               REGION "BUTTON 3"
                   #btnActivateInt[3] := #btn3Activate;
                   #btnModeInt[3] := #btn3Mode;
                   #btnGroup[3] := #btn3Group;
                   #btnClrOn1Int[3] := #btn3ColorOn1;
                   #btnClrOn2Int[3] := #btn3ColorOn2;
                   #btnClrOffInt[3] := #btn3ColorOff;
               END_REGION

               REGION "BUTTON 4"
                   #btnActivateInt[4] := #btn4Activate;
                   #btnModeInt[4] := #btn4Mode;
                   #btnGroup[4] := #btn4Group;
                   #btnClrOn1Int[4] := #btn4ColorOn1;
                   #btnClrOn2Int[4] := #btn4ColorOn2;
                   #btnClrOffInt[4] := #btn4ColorOff;
               END_REGION

               REGION "BUTTON 5"
                   #btnActivateInt[5] := #btn5Activate;
                   #btnModeInt[5] := #btn5Mode;
                   #btnGroup[5] := #btn5Group;
                   #btnClrOn1Int[5] := #btn5ColorOn1;
                   #btnClrOn2Int[5] := #btn5ColorOn2;
                   #btnClrOffInt[5] := #btn5ColorOff;
               END_REGION

               REGION "BUTTON 6"
                   #btnActivateInt[6] := #btn6Activate;
                   #btnModeInt[6] := #btn6Mode;
                   #btnGroup[6] := #btn6Group;
                   #btnClrOn1Int[6] := #btn6ColorOn1;
                   #btnClrOn2Int[6] := #btn6ColorOn2;
                   #btnClrOffInt[6] := #btn6ColorOff;
               END_REGION

               REGION "BUTTON 7"
                   #btnActivateInt[7] := #btn7Activate;
                   #btnModeInt[7] := #btn7Mode;
                   #btnGroup[7] := #btn7Group;
                   #btnClrOn1Int[7] := #btn7ColorOn1;
                   #btnClrOn2Int[7] := #btn7ColorOn2;
                   #btnClrOffInt[7] := #btn7ColorOff;
               END_REGION

           END_REGION

           REGION "RECOLOR BUTTON MASKS"
               FOR #i1 := 0 TO 7 DO

                   REGION "ON COLOR 1"
                       IF (#btnClrOn1Int[#i1] = 'red') THEN
                           #btnClrMskOn1Int[#i1] := SHL(IN := #btnMskRed, N := INT_TO_ULINT(#i1));
                       ELSIF (#btnClrOn1Int[#i1] = 'green') THEN
                           #btnClrMskOn1Int[#i1] := SHL(IN := #btnMskGreen, N := INT_TO_ULINT(#i1));
                       ELSIF (#btnClrOn1Int[#i1] = 'blue') THEN
                           #btnClrMskOn1Int[#i1] := SHL(IN := #btnMskBlue, N := INT_TO_ULINT(#i1));
                       ELSIF (#btnClrOn1Int[#i1] = 'yellow') THEN
                           #btnClrMskOn1Int[#i1] := SHL(IN := #btnMskYellow, N := INT_TO_ULINT(#i1));
                       ELSIF (#btnClrOn1Int[#i1] = 'white') THEN
                           #btnClrMskOn1Int[#i1] := SHL(IN := #btnMskWhite, N := INT_TO_ULINT(#i1));
                       ELSIF (#btnClrOn1Int[#i1] = 'off') THEN
                           #btnClrMskOn1Int[#i1] := 0;
                       END_IF;
                   END_REGION

                   REGION "ON COLOR 2"
                       IF (#btnClrOn2Int[#i1] = 'red') THEN
                           #btnClrMskOn2Int[#i1] := SHL(IN := #btnMskRed, N := INT_TO_ULINT(#i1));
                       ELSIF (#btnClrOn2Int[#i1] = 'green') THEN
                           #btnClrMskOn2Int[#i1] := SHL(IN := #btnMskGreen, N := INT_TO_ULINT(#i1));
                       ELSIF (#btnClrOn2Int[#i1] = 'blue') THEN
                           #btnClrMskOn2Int[#i1] := SHL(IN := #btnMskBlue, N := INT_TO_ULINT(#i1));
                       ELSIF (#btnClrOn2Int[#i1] = 'yellow') THEN
                           #btnClrMskOn2Int[#i1] := SHL(IN := #btnMskYellow, N := INT_TO_ULINT(#i1));
                       ELSIF (#btnClrOn2Int[#i1] = 'white') THEN
                           #btnClrMskOn2Int[#i1] := SHL(IN := #btnMskWhite, N := INT_TO_ULINT(#i1));
                       ELSIF (#btnClrOn2Int[#i1] = 'off') THEN
                           #btnClrMskOn2Int[#i1] := 0;
                       END_IF;
                   END_REGION

                   REGION "OFF COLOR"
                       IF (#btnClrOffInt[#i1] = 'red') THEN
                           #btnClrMskOffInt[#i1] := SHL(IN := #btnMskRed, N := INT_TO_ULINT(#i1));
                       ELSIF (#btnClrOffInt[#i1] = 'green') THEN
                           #btnClrMskOffInt[#i1] := SHL(IN := #btnMskGreen, N := INT_TO_ULINT(#i1));
                       ELSIF (#btnClrOffInt[#i1] = 'blue') THEN
                           #btnClrMskOffInt[#i1] := SHL(IN := #btnMskBlue, N := INT_TO_ULINT(#i1));
                       ELSIF (#btnClrOffInt[#i1] = 'yellow') THEN
                           #btnClrMskOffInt[#i1] := SHL(IN := #btnMskYellow, N := INT_TO_ULINT(#i1));
                       ELSIF (#btnClrOffInt[#i1] = 'white') THEN
                           #btnClrMskOffInt[#i1] := SHL(IN := #btnMskWhite, N := INT_TO_ULINT(#i1));
                       ELSIF (#btnClrOffInt[#i1] = 'off') THEN
                           #btnClrMskOffInt[#i1] := 0;
                       END_IF;
                   END_REGION

               END_FOR;
           END_REGION

       END_IF;
   END_REGION

   REGION "HART INIT"
       IF #hardInit THEN
           FOR #i1 := 0 TO 7 DO
               #btnStateArrayInt[#i1] := FALSE;
           END_FOR;
       END_IF;
   END_REGION


   REGION "TRANFER PARAMETERS TO ARRAYS"
       // raw pb data
       #btnInInt := #btnIn;
       // flashing modes
       #btnFlashInt[0] := #btn0Flash;
       #btnFlashInt[1] := #btn1Flash;
       #btnFlashInt[2] := #btn2Flash;
       #btnFlashInt[3] := #btn3Flash;
       #btnFlashInt[4] := #btn4Flash;
       #btnFlashInt[5] := #btn5Flash;
       #btnFlashInt[6] := #btn6Flash;
       #btnFlashInt[7] := #btn7Flash;
   END_REGION

   REGION "EVALUATE BUTTONS"
       FOR #i1 := 0 TO 7 DO

           REGION "TRANSFER BUTTON PRESSES TO ARRAY"
               #btnEval := SHR(IN := #btnInInt, N := INT_TO_ULINT(#i1));
               #btnInArrayNew[#i1] := #btnEval.%X0;
               #btnEval := b#16#0;
           END_REGION

           REGION "SET BUTTON STATE"

               REGION "BUTTON ACTIVE"
                   IF #btnActivateInt[#i1] THEN

                       REGION "MAINTAINED"
                           IF #btnModeInt[#i1] THEN

                               REGION "RISING EDGE OF PRESS"
                                   IF #btnInArrayNew[#i1] AND NOT #btnInArrayOld[#i1] THEN

                                       REGION "CHECK FOR GROUP MEMBERSHIP"
                                           FOR #i2 := 0 TO 7 DO

                                               REGION "NOT IN NULL GROUP"
                                                   IF (#btnGroup[#i2] <> 0) THEN

                                                       REGION "SKIP SELF"
                                                           IF (#i2 <> #i1) THEN

                                                               REGION "GROUPS MATCH"
                                                                   IF #btnGroup[#i1] = #btnGroup[#i2] THEN
                                                                       REGION "DEACTIVATE OTHER GROUP MEMBERS"
                                                                           #btnStateArrayInt[#i2] := FALSE;
                                                                       END_REGION

                                                                   END_IF;
                                                               END_REGION

                                                           END_IF;
                                                       END_REGION

                                                   END_IF;
                                               END_REGION

                                           END_FOR;
                                       END_REGION

                                       REGION "TOGGLE STATE"
                                           #btnStateArrayInt[#i1] := NOT #btnStateArrayInt[#i1];
                                       END_REGION

                                   END_IF;
                               END_REGION

                           END_IF;
                       END_REGION

                       REGION "MOMENTARY"
                           IF NOT #btnModeInt[#i1] THEN
                               #btnStateArrayInt[#i1] := #btnInArrayNew[#i1];
                           END_IF;
                       END_REGION

                   END_IF;
               END_REGION

               REGION "BUTTON INACTIVE"
                   IF NOT #btnActivateInt[#i1] THEN
                       #btnStateArrayInt[#i1] := FALSE;
                   END_IF;
               END_REGION

           END_REGION

           REGION "ANIMATE BUTTONS"

               REGION "BUTTON ON FLASH BIT OFF"
                   IF #btnStateArrayInt[#i1] AND NOT #btnFlashInt[#i1] THEN
                       #btnColors := #btnColors AND ROL(IN := #btnMskBlack, N := INT_TO_ULINT(#i1));
                       #btnColors := #btnColors OR #btnClrMskOn1Int[#i1];
                   END_IF;
               END_REGION

               REGION "BUTTON ON FLASH BIT ON"
                   IF #btnStateArrayInt[#i1] AND #btnFlashInt[#i1] THEN
                       #btnColors := #btnColors AND ROL(IN := #btnMskBlack, N := INT_TO_ULINT(#i1));
                       #btnColors := #btnColors OR #btnClrMskOn2Int[#i1];
                   END_IF;
               END_REGION

               REGION "BUTTON OFF"
                   IF NOT #btnStateArrayInt[#i1] THEN
                       #btnColors := #btnColors AND ROL(IN := #btnMskBlack, N := INT_TO_ULINT(#i1));
                       #btnColors := #btnColors OR #btnClrMskOffInt[#i1];
                   END_IF;
               END_REGION

           END_REGION

       END_FOR;
   END_REGION

   REGION "CHANGE DETECTION"
       #btnInArrayOld := #btnInArrayNew;
   END_REGION

   REGION "OUTPUT"
       #btnColorsOut := #btnColors;
       #btnStatesOut := #btnStateArrayInt;
   END_REGION
END_FUNCTION_BLOCK

FUNCTION "Physical to Global" : Void   // FC1, LAD
{ S7_Optimized_Access := 'TRUE' }
VERSION : 0.1
   VAR_IN_OUT
      stations : "Stations";
   END_VAR
   VAR_TEMP
      i : Int;
      kp8In : DWord;
   END_VAR
BEGIN

REGION Network 1 (SCL): MAIN LOOP
   FOR #i := 0 TO "stnCount" DO

       CASE #i OF
           "VOLVO 16 01":
               #kp8In := "VOLVO 16 01 KP8 In";
           "VOLVO 16 02":
               #kp8In := "VOLVO 16 02 KP8 In";
           "VOLVO 16 03":
               #kp8In := "VOLVO 16 03 KP8 In";
           "VOLVO 16 04":
               #kp8In := "VOLVO 16 04 KP8 In";
           "VOLVO 16 05":
               #kp8In := "VOLVO 16 05 KP8 In";
           "VOLVO 16 06":
               #kp8In := "VOLVO 16 06 KP8 In";
           "VOLVO 16 07":
               #kp8In := "VOLVO 16 07 KP8 In";
           "VOLVO 16 08":
               #kp8In := "VOLVO 16 08 KP8 In";
           "VOLVO 16 09":
               #kp8In := "VOLVO 16 09 KP8 In";
           "VOLVO 16 10":
               #kp8In := "VOLVO 16 10 KP8 In";
           "VOLVO 16 11":
               #kp8In := "VOLVO 16 11 KP8 In";
           "CHM 01":
               #kp8In := "CHM 01 KP8 In";
           "CHM 02":
               #kp8In := "CHM 02 KP8 In";
           "CHM 03":
               #kp8In := "CHM 03 KP8 In";
           "CHM 04":
               #kp8In := "CHM 04 KP8 In";
           "CHM 05":
               #kp8In := "CHM 05 KP8 In";
           "CDO 01":
               #kp8In := "CDO 01 KP8 In";
           "CDO 02":
               #kp8In := "CDO 02 KP8 In";
           "CDO 03":
               #kp8In := "CDO 03 KP8 In";
           "BFL 01":
               #kp8In := "BFL 01 KP8 In";
           "BFL 02":
               #kp8In := "BFL 02 KP8 In";
           "BFL 03":
               #kp8In := "BFL 03 KP8 In";
           "LGS 01":
               #kp8In := "LGS 01 KP8 In";
           "LGS 02":
               #kp8In := "LGS 02 KP8 In";

       END_CASE;

       #stations.me[#i].kp8In := #kp8In.%B3;

   END_FOR;
END_REGION
END_FUNCTION

FUNCTION "Time to WString" : WString   // FC2, SCL
{ S7_Optimized_Access := 'TRUE' }
VERSION : 0.1
   VAR_INPUT
      "Time" : Time;
   END_VAR
   VAR_TEMP
      "Time as DInt" : DInt;
      "Hours 10s Place" : DInt;
      "Hours 1s Place" : DInt;
      "Minutes 10s Place" : DInt;
      "Minutes 1s Place" : DInt;
      "Seconds 10s Place" : DInt;
      "Seconds 1s Place" : DInt;
      "Time Elements" : Array[0..4] of WString;
      Length : Int;
      "String Box" : WString;
      "DInt Box" : DInt;
   END_VAR
   VAR CONSTANT
      "Milliseconds per 10 Hours" : DInt := 36000000;
      "Milliseconds per Hour" : DInt := 3600000;
      "Milliseconds per 10 Minutes" : DInt := 600000;
      "Milliseconds per Minute" : DInt := 60000;
      "Milliseconds per 10 Seconds" : DInt := 10000;
      "Milliseconds per Second" : DInt := 1000;
   END_VAR
BEGIN
   REGION GET INPUT
       #"Time as DInt" := #Time;
   END_REGION

   REGION CONVERT TIME INTO INDIVIDUAL PLACE VALUES
       #"Minutes 10s Place" := #"Time as DInt" / #"Milliseconds per 10 Minutes";
       #"Minutes 1s Place" := (#"Time as DInt" / #"Milliseconds per Minute") MOD 10;
       #"Seconds 10s Place" := (#"Time as DInt" MOD #"Milliseconds per Minute") / #"Milliseconds per 10 Seconds";
       #"Seconds 1s Place" := (#"Time as DInt" / #"Milliseconds per Second") MOD 10;
   END_REGION

   REGION "ADD SIGN"
       #"Time Elements"[0] := wstring#'';
       IF #"Minutes 10s Place" < 0 OR
           #"Minutes 1s Place" < 0 OR
           #"Seconds 10s Place" < 0 OR
           #"Seconds 1s Place" < 0 THEN
            #"Time Elements"[0] := wstring#'-';
       END_IF;
   END_REGION

   REGION CONVERT PLACE VALUES INTO COMPONENT STRINGS
       // MINUTES
       #"DInt Box" := #"Minutes 10s Place" * 10 + #"Minutes 1s Place";
       #"String Box" := DINT_TO_WSTRING(IN := #"DInt Box");
       #"String Box" := "Strip Sign"("WString":=#"String Box");
       #"String Box" := "Add Leading"("Leading Character" := WCHAR#'0',
                                      "Desired Length" := 2,
                                      "String" := #"String Box");
       #"Time Elements"[1] := #"String Box";
       // COLON
       #"Time Elements"[2] := WSTRING#':';
       // SECONDS
       #"DInt Box" := #"Seconds 10s Place" * 10 + #"Seconds 1s Place";
       #"String Box" := DINT_TO_WSTRING(IN := #"DInt Box");
       #"String Box" := "Strip Sign"("WString":=#"String Box");
       #"String Box" := "Add Leading"("Leading Character" := WCHAR#'0',
                                      "Desired Length" := 2,
                                      "String" := #"String Box");
       #"Time Elements"[3] := #"String Box";
   END_REGION


   REGION RETURN VALUE
       #"Time to WString" := CONCAT_WSTRING(IN1 := #"Time Elements"[0],
                                            IN2 := #"Time Elements"[1],
                                            IN3 := #"Time Elements"[2],
                                            IN4 := #"Time Elements"[3]);
   END_REGION
END_FUNCTION

FUNCTION "Strip Sign" : WString   // FC3, SCL
{ S7_Optimized_Access := 'TRUE' }
VERSION : 0.1
   VAR_INPUT
      WString : WString;
   END_VAR
   VAR_TEMP
      Length : Int;
      "String Box" : WString;
      "Test Character" : WString;
   END_VAR
   VAR CONSTANT
      "+" : WChar := WCHAR#'+';
      "-" : WChar := WCHAR#'-';
   END_VAR
BEGIN
   #"String Box" := #WString;
   #"Test Character" := LEFT_WSTRING(IN := #"String Box",
                                     L := 1);
   IF #"Test Character" = #"+" OR #"Test Character" = #"-" THEN
       #Length := LEN(#"String Box");
       #"String Box" := RIGHT_WSTRING(IN := #"String Box", L := #Length - 1);

   END_IF;
   #"Strip Sign" := #"String Box";
END_FUNCTION

FUNCTION "Add Leading" : WString   // FC4, SCL
{ S7_Optimized_Access := 'TRUE' }
VERSION : 0.1
   VAR_INPUT
      "Leading Character" : WChar;
      "Desired Length" : USInt;
      "String" : WString;
   END_VAR
   VAR_TEMP
      Length : Int;
      "String Box" : WString;
      Constant : WString;
   END_VAR
BEGIN
   #"String Box" := #String;
   #Length := LEN(#"String Box");

   WHILE #Length < #"Desired Length" DO
       #"String Box" := CONCAT_WSTRING(IN1 := #"Leading Character",
                                       IN2 := #"String Box");
       #Length := LEN(#"String Box");
   END_WHILE;

   #"Add Leading" := #"String Box";
END_FUNCTION

FUNCTION "Global to Physical" : Void   // FC5, LAD
{ S7_Optimized_Access := 'TRUE' }
VERSION : 0.1
   VAR_IN_OUT
      stations : "Stations";
   END_VAR
   VAR_TEMP
      i : Int;
      j : Int;
      IO : DWord;
      "KP8 In" : DWord;
      "KP8 Out" : DWord;
      Card : Int;
      stnCount : Int;
   END_VAR
   VAR CONSTANT
      "VOLVO 16 01" : Int := 0;
      "VOLVO 16 02" : Int := 1;
      "VOLVO 16 03" : Int := 2;
      "VOLVO 16 04" : Int := 3;
      "VOLVO 16 05" : Int := 4;
      "VOLVO 16 06" : Int := 5;
      "VOLVO 16 07" : Int := 6;
      "VOLVO 16 08" : Int := 7;
      "VOLVO 16 09" : Int := 8;
      "VOLVO 16 10" : Int := 9;
      "VOLVO 16 11" : Int := 10;
      "CHM 01" : Int := 11;
      "CHM 02" : Int := 12;
      "CHM 03" : Int := 13;
      "CHM 04" : Int := 14;
      "CHM 05" : Int := 15;
      "CDO 01" : Int := 16;
      "CDO 02" : Int := 17;
      "CDO 03" : Int := 18;
      "BFL 01" : Int := 19;
      "BFL 02" : Int := 20;
      "BFL 03" : Int := 21;
      "LGS 01" : Int := 22;
      "LGS 02" : Int := 23;
   END_VAR
BEGIN

REGION Network 1: ARRAY LIMIT FOR STATION COUNT
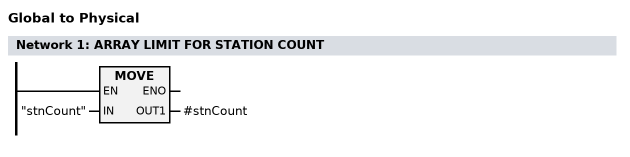
   RUNG wire#powerrail
      Move(in := "stnCount", out1 => #stnCount)
   END_RUNG
   // the same network as SCL:
   #stnCount := "stnCount";
END_REGION

REGION Network 2 (SCL): MAIN LOOP
   FOR #i := 0 TO #stnCount DO

       #IO := #stations.me[#i].stackLightOut;
       #"KP8 Out" := #stations.me[#i].kp8Out;

       CASE #i OF
           #"VOLVO 16 01":
               "VOLVO 16 01 IO" := #IO;
               "VOLVO 16 01 KP8 Out" := #"KP8 Out";
           #"VOLVO 16 02":
               "VOLVO 16 02 IO" := #IO;
               "VOLVO 16 02 KP8 Out" := #"KP8 Out";
           #"VOLVO 16 03":
               "VOLVO 16 03 IO" := #IO;
               "VOLVO 16 03 KP8 Out" := #"KP8 Out";
           #"VOLVO 16 04":
               "VOLVO 16 04 IO" := #IO;
               "VOLVO 16 04 KP8 Out" := #"KP8 Out";
           #"VOLVO 16 05":
               "VOLVO 16 05 IO" := #IO;
               "VOLVO 16 05 KP8 Out" := #"KP8 Out";
           #"VOLVO 16 06":
               "VOLVO 16 06 IO" := #IO;
               "VOLVO 16 06 KP8 Out" := #"KP8 Out";
           #"VOLVO 16 07":
               "VOLVO 16 07 IO" := #IO;
               "VOLVO 16 07 KP8 Out" := #"KP8 Out";
           #"VOLVO 16 08":
               "VOLVO 16 08 IO" := #IO;
               "VOLVO 16 08 KP8 Out" := #"KP8 Out";
           #"VOLVO 16 09":
               "VOLVO 16 09 IO" := #IO;
               "VOLVO 16 09 KP8 Out" := #"KP8 Out";
           #"VOLVO 16 10":
               "VOLVO 16 10 IO" := #IO;
               "VOLVO 16 10 KP8 Out" := #"KP8 Out";
           #"VOLVO 16 11":
               "VOLVO 16 11 IO" := #IO;
               "VOLVO 16 11 KP8 Out" := #"KP8 Out";
           #"CHM 01":
               "CHM 01 IO" := #IO;
               "CHM 01 KP8 Out" := #"KP8 Out";
           #"CHM 02":
               "CHM 02 IO" := #IO;
               "CHM 02 KP8 Out" := #"KP8 Out";
           #"CHM 03":
               "CHM 03 IO" := #IO;
               "CHM 03 KP8 Out" := #"KP8 Out";
           #"CHM 04":
               "CHM 04 IO" := #IO;
               "CHM 04 KP8 Out" := #"KP8 Out";
           #"CHM 05":
               "CHM 05 IO" := #IO;
               "CHM 05 KP8 Out" := #"KP8 Out";
           #"CDO 01":
               "CDO 01 IO" := #IO;
               "CDO 01 KP8 Out" := #"KP8 Out";
           #"CDO 02":
               "CDO 02 IO" := #IO;
               "CDO 02 KP8 Out" := #"KP8 Out";
           #"CDO 03":
               "CDO 03 IO" := #IO;
               "CDO 03 KP8 Out" := #"KP8 Out";
           #"BFL 01":
               "BFL 01 IO" := #IO;
               "BFL 01 KP8 Out" := #"KP8 Out";
           #"BFL 02":
               "BFL 02 IO" := #IO;
               "BFL 02 KP8 Out" := #"KP8 Out";
           #"BFL 03":
               "BFL 03 IO" := #IO;
               "BFL 03 KP8 Out" := #"KP8 Out";
           #"LGS 01":
               "LGS 01 IO" := #IO;
               "LGS 01 KP8 Out" := #"KP8 Out";
           #"LGS 02":
               "LGS 02 IO" := #IO;
               "LGS 02 KP8 Out" := #"KP8 Out";

       END_CASE;

   END_FOR;
END_REGION
END_FUNCTION

FUNCTION "Select Stations" : Void   // FC6, SCL
{ S7_Optimized_Access := 'TRUE' }
VERSION : 0.1
   VAR_INPUT
      mode : Bool;   // TRUE = select; FALSE = deselect
   END_VAR
   VAR_IN_OUT
      stations : "Stations";
   END_VAR
   VAR_TEMP
      i : Int;
      stnCount : Int;
   END_VAR
   VAR CONSTANT
      stationCount : Int := 22;
   END_VAR
BEGIN
   REGION "GET STATION COUNT"
       #stnCount := "stnCount";
   END_REGION

   REGION "SELECT STATIONS"
       FOR #i := 0 TO #stnCount DO
           #stations.me[#i].settings.selected := #mode;
       END_FOR;
   END_REGION
END_FUNCTION

FUNCTION "Dark Mode" : Void   // FC7, SCL
{ S7_Optimized_Access := 'TRUE' }
VERSION : 0.1
   VAR_IN_OUT
      animate : USInt;
   END_VAR
   VAR_TEMP
      ani : USInt;
   END_VAR
   VAR CONSTANT
      redFlashing : USInt := 12;
      invisible : USInt := 255;
      darkMode : USInt := 1;
      disabled : USInt := 254;
   END_VAR
BEGIN
   REGION "COPY TO LOCAL"
       #ani := #animate;
   END_REGION


   REGION "APPLY DARK MODE"
       CASE #ani OF
           #redFlashing, #invisible, 0, #disabled:
               #ani := #ani;
           ELSE
               #ani += #darkMode;
       END_CASE;
   END_REGION


   REGION "OUTPUT"
       #animate := #ani;
   END_REGION
END_FUNCTION

FUNCTION "Select Buttons" : Void   // FC8, SCL
{ S7_Optimized_Access := 'TRUE' }
VERSION : 0.1
   VAR_INPUT
      mode : Bool;   // TRUE = select; FALSE = deselect
   END_VAR
   VAR_IN_OUT
      stations : "Stations";
   END_VAR
   VAR_TEMP
      btnCount : Int;
      i : Int;
      j : Int;
      selected : Bool;
      stnCount : Int;
   END_VAR
   VAR CONSTANT
      buttonCount : Int := 5;
   END_VAR
BEGIN
   REGION "COPY TO LOCAL"
       #btnCount := "ptsPerStn";
       #stnCount := "stnCount";
   END_REGION

   REGION "SELECT BUTTONS"
       FOR #i := 0 TO #stnCount DO

           REGION "SELCT ALL BUTTONS ON SELECTED STATION"
               #selected := #stations.me[#i].settings.selected;
               IF #selected THEN

                   REGION "LOOP THROUGH BUTTONS"
                       FOR #j := 0 TO #btnCount DO
                           #stations.me[#i].settings.btnSelection[#j] := #mode;
                       END_FOR;
                   END_REGION

               END_IF;
           END_REGION

       END_FOR;
   END_REGION
END_FUNCTION

FUNCTION "Animate Bool" : USInt   // FC9, SCL
{ S7_Optimized_Access := 'TRUE' }
VERSION : 0.1
   VAR_INPUT
      colorTrue : USInt;
      colorFalse : USInt;
      evalSignal : Bool;
   END_VAR
   VAR_TEMP
      animate : USInt;
   END_VAR
BEGIN
   REGION "FALSE COLOR"
       IF NOT #evalSignal THEN
           #animate := #colorFalse;
       END_IF;
   END_REGION

   REGION "TRUE COLOR"
       IF #evalSignal THEN
           #animate := #colorTrue;
       END_IF;
   END_REGION

   REGION "FUNCTION RETURN"
       #"Animate Bool" := #animate;
   END_REGION
END_FUNCTION

FUNCTION "WString to Time" : Time   // FC10, SCL
{ S7_Optimized_Access := 'TRUE' }
VERSION : 0.1
   VAR_INPUT
      WString : WString;
   END_VAR
   VAR_TEMP
      Count : UInt;
      "DInt Box" : DInt;
      "String Box" : WString [5];
      "Time Box" : Time;
      "WChar Array" : Array[0..4] of WChar;
   END_VAR
   VAR CONSTANT
      "ms/(10 hr)" : DInt := 36000000;
      "ms/hr" : DInt := 3600000;
      "ms/(10 min)" : DInt := 600000;
      "ms/min" : DInt := 60000;
      "ms/(10 sec)" : DInt := 10000;
      "ms/sec" : DInt := 1000;
   END_VAR
BEGIN
   REGION EXPLODE INPUT

       #"String Box" := #WString;
       IF #"String Box" = WSTRING#'' THEN
           #"String Box" := WSTRING#'00:00';
       END_IF;

       Strg_TO_Chars(Strg := #"String Box",
                     pChars := 0,
                     Cnt => #Count,
                     Chars := #"WChar Array");

   END_REGION

   REGION CONVERT ARRAY ELEMENTS TO TIME

       // 10S OF MINUTES
       #"DInt Box" := WCHAR_TO_DINT(IN := #"WChar Array"[0]) - 16#30;
       #"Time Box" := #"Time Box" + #"DInt Box" * #"ms/(10 min)";

       // MINUTES
       #"DInt Box" := WCHAR_TO_DINT(IN := #"WChar Array"[1]) - 16#30;
       #"Time Box" := #"Time Box" + #"DInt Box" * #"ms/min";

       // 10S OF SECONDS
       #"DInt Box" := WCHAR_TO_DINT(IN := #"WChar Array"[3]) - 16#30;
       #"Time Box" := #"Time Box" + #"DInt Box" * #"ms/(10 sec)";

       // SECONDS
       #"DInt Box" := WCHAR_TO_DINT(IN := #"WChar Array"[4]) - 16#30;
       #"Time Box" := #"Time Box" + #"DInt Box" * #"ms/sec";

   END_REGION


   REGION RETURN VALUE

       #"WString to Time" := #"Time Box";

   END_REGION
END_FUNCTION

FUNCTION "Get Part Call Row Number" : Int   // FC11, SCL
{ S7_Optimized_Access := 'TRUE' }
VERSION : 0.1
   VAR_IN_OUT
      partCall : "Part Call Screen";
   END_VAR
   VAR_TEMP
      hmiRows : Int;
      i : Int;
      selectedRow : Int;
   END_VAR
BEGIN
   REGION "GET NUMBER OF HMI ROWS"
       #hmiRows := "partReqHmiRowCount";
   END_REGION

   REGION "LOOP THROUGH HMI ROWS
       FOR #i := 0 TO #hmiRows DO

           REGION "FIND SELECTED ROW"
               IF #partCall.row[#i].pbSelection.actuate THEN
                   // selected row as int
                   #selectedRow := #i + 1;
                   EXIT;
               END_IF;
           END_REGION

       END_FOR;
   END_REGION

   REGION "RETURN ROW NUMBER"
       #"Get Part Call Row Number" := #selectedRow;
   END_REGION
END_FUNCTION

FUNCTION "Address to Station and Button" : Void   // FC12, SCL
{ S7_Optimized_Access := 'TRUE' }
VERSION : 0.1
   VAR_INPUT
      address : UInt;
   END_VAR
   VAR_OUTPUT
      station : UInt;
      button : UInt;
   END_VAR
BEGIN
   #station := #address / 10;
   #button := #address MOD 10;
END_FUNCTION

FUNCTION "WString Timer to Real" : Real   // FC13, SCL
{ S7_Optimized_Access := 'TRUE' }
VERSION : 0.1
   VAR_INPUT
      wstring : WString;
   END_VAR
   VAR CONSTANT
      msPerSec : Real := 1000.0;
   END_VAR
BEGIN
   #"WString Timer to Real" := DINT_TO_REAL(TIME_TO_DINT("WString to Time"(#wstring))) / #msPerSec;
END_FUNCTION

FUNCTION "Real to WString Timer" : WString   // FC14, SCL
{ S7_Optimized_Access := 'TRUE' }
VERSION : 0.1
   VAR_INPUT
      realVal : Real;
   END_VAR
   VAR CONSTANT
      msPerSec : Real := 1000.0;
   END_VAR
BEGIN
   #"Real to WString Timer" := "Time to WString"(DINT_TO_TIME(REAL_TO_DINT(#realVal * #msPerSec)));
END_FUNCTION

FUNCTION "Populate Dropzone IO Field" : WString   // FC15, SCL
{ S7_Optimized_Access := 'TRUE' }
VERSION : 0.1
   VAR_INPUT
      dzAsInt : USInt;
   END_VAR
BEGIN
   #"Populate Dropzone IO Field" := "Strip Sign"(USINT_TO_WSTRING(#dzAsInt));
END_FUNCTION

FUNCTION "Get Station Selection Number" : Void   // FC16, SCL
{ S7_Optimized_Access := 'TRUE' }
VERSION : 0.1
   VAR_INPUT
      next : Bool;   // 'next' or 'prev'
      prev : Bool;
      stations : "Stations";
   END_VAR
   VAR_IN_OUT
      selStnNumber : Int;
   END_VAR
   VAR_TEMP
      i : Int;
      stnCount : Int;
      stnSelected : Bool;
   END_VAR
BEGIN
   REGION "COPY TO LOCAL"
       #stnCount := "stnCount";
   END_REGION

   REGION "INITIALIZE INDEX"
       #i := #selStnNumber;
   END_REGION

   REGION "PREVIOUS MODE"

       REGION "DECREMENT"
           IF #prev THEN
               #i -= 1;
           END_IF;
       END_REGION

       REGION "LOW LIMIT ROLLOVER"
           IF #i < 0 THEN
               #i := #stnCount;
           END_IF;
       END_REGION

   END_REGION

   REGION "NEXT MODE"

       REGION "INCREMENT"
           IF #next THEN
               #i += 1;
           END_IF;
       END_REGION

       REGION "HIGH LIMIT ROLLOVER"
           IF #i > #stnCount THEN
               #i := 0;
           END_IF;
       END_REGION

   END_REGION

   REGION "COPY TO LOCAL"
       #stnSelected := #stations.me[#i].settings.selected;
   END_REGION

   REGION "FIND NEXT SELECTED STATION"
       WHILE NOT #stnSelected DO

           REGION "PREVIOUS MODE"

               REGION "DECREMENT"
                   IF #prev THEN
                       #i -= 1;
                   END_IF;
               END_REGION

               REGION "LOW LIMIT ROLLOVER"
                   IF #i < 0 THEN
                       #i := #stnCount;
                   END_IF;
               END_REGION

           END_REGION

           REGION "NEXT MODE"

               REGION "INCREMENT"
                   IF #next THEN
                       #i += 1;
                   END_IF;
               END_REGION

               REGION "HIGH LIMIT ROLLOVER"
                   IF #i > #stnCount THEN
                       #i := 0;
                   END_IF;
               END_REGION

           END_REGION

           REGION "SAVE WHILE CONDITION"
               #stnSelected := #stations.me[#i].settings.selected;
           END_REGION

       END_WHILE;
   END_REGION

   REGION "RETURN VALUE"
       #selStnNumber := #i;
   END_REGION
END_FUNCTION

FUNCTION "Populate Button Details" : Void   // FC17, SCL
{ S7_Optimized_Access := 'TRUE' }
VERSION : 0.1
   VAR_INPUT
      selStnNumber : Int;
      stations : "Stations";
   END_VAR
   VAR_IN_OUT
      settings : "Settings";
   END_VAR
   VAR_TEMP
      btnCount : Int;
      i : Int;
      partNumber : WString;
      pBtn : Int;
      timerWS : WString;
   END_VAR
BEGIN
   REGION "COPY TO LOCAL"
       #btnCount := "ptsPerStn";
   END_REGION

   REGION "FOR EACH BUTTON"
       FOR #i := 0 TO #btnCount DO

           REGION "CALCULATE BUTTON POINTER"
               IF #i MOD 2 = 0 THEN
                   #pBtn := 7 - #i / 2;
               END_IF;
               IF #i MOD 2 <> 0 THEN
                   #pBtn := 3 - #i / 2;
               END_IF;
           END_REGION

           REGION "BUTTON LABEL"
               #settings.viewingStation.btns[#i].label.value := "Strip Sign"(INT_TO_WSTRING(#i + 1));
           END_REGION

           REGION "ALLOTTED TIME"
               #timerWS := "Real to WString Timer"(#stations.me[#selStnNumber].presetTime.allotted[#pBtn]);
               #settings.viewingStation.btns[#i].alloted.value := #timerWS;
           END_REGION

           REGION "CRITICAL TIME"
               #timerWS := "Real to WString Timer"(#stations.me[#selStnNumber].presetTime.critical[#pBtn]);
               #settings.viewingStation.btns[#i].critical.value := #timerWS;
           END_REGION

           REGION "PART NUMBER"
               #partNumber := #stations.me[#selStnNumber].partNumbers[#pBtn];
               #settings.viewingStation.btns[#i].partNumber.value := #partNumber;
           END_REGION

       END_FOR;
   END_REGION
END_FUNCTION

FUNCTION "Assign Station Parameters" : Void   // FC18, SCL
{ S7_Optimized_Access := 'TRUE' }
VERSION : 0.1
   VAR_IN_OUT
      settings : "Settings";
      stations : "Stations";
   END_VAR
   VAR_TEMP
      dzEntered : Bool;
      dzLabel : WString;
      i : Int;
      lineEntered : Bool;
      lineLabel : WString;
      stnCount : Int;
      stnSelected : Bool;
   END_VAR
BEGIN
   REGION "COPY TO LOCAL"    
       #dzEntered := #settings.viewingStation.dzData.inputFinished;
       #lineEntered := #settings.viewingStation.lineData.inputFinished;
       #stnCount := "stnCount";
   END_REGION

   REGION "ON PARAMETER ENTRY"
       IF #dzEntered OR #lineEntered THEN

           REGION "TURN OFF THE LIGHTS"
               #settings.viewingStation.dzData.inputFinished := FALSE;
               #settings.viewingStation.lineData.inputFinished := FALSE;
           END_REGION

           REGION "FOR EACH STATION"
               FOR #i := 0 TO #stnCount DO

                   REGION "COPY TO LOCAL"
                       #stnSelected := #stations.me[#i].settings.selected;
                   END_REGION

                   REGION "ON SELECTED STATION"
                       IF #stnSelected THEN

                           REGION "ON DROP ZONE INPUT"
                               IF #dzEntered THEN

                                   REGION "GET FROM HMI"
                                       #dzLabel := #settings.viewingStation.dzData.value;
                                   END_REGION

                                   REGION "WRITE TO STATION PARAMETER"
                                       #stations.me[#i].dropZone := WSTRING_TO_USINT(#dzLabel);
                                   END_REGION

                               END_IF;
                           END_REGION

                           REGION "ON LINE LABEL INPUT"
                               IF #lineEntered THEN

                                   REGION "GET FROM HMI"
                                       #lineLabel := #settings.viewingStation.lineData.value;
                                   END_REGION

                                   REGION "WRITE TO STATION PARAMETER"
                                       #stations.me[#i].line := #lineLabel;
                                   END_REGION

                               END_IF;
                           END_REGION

                       END_IF;
                   END_REGION

               END_FOR;
           END_REGION

       END_IF;
   END_REGION
END_FUNCTION

FUNCTION "Animate Button Details" : Void   // FC19, SCL
{ S7_Optimized_Access := 'TRUE' }
VERSION : 0.1
   VAR_INPUT
      stations : "Stations";
   END_VAR
   VAR_IN_OUT
      settings : "Settings";
   END_VAR
   VAR_TEMP
      animate : USInt;
      btnCount : Int;
      btnSelected : Bool;
      deselected : USInt;
      i : Int;
      invisible : USInt;
      pBtn : Int;
      selected : USInt;
      selStnCount : Int;
      selStnNumber : Int;
   END_VAR
BEGIN
   REGION "COPY TO LOCAL"
       #btnCount := "ptsPerStn";
       #deselected := "BgGray";
       #invisible := "invisible";
       #selected := "BgLTe";
       #selStnCount := #settings.#stations.selCount;
       #selStnNumber := #settings.stations.selNumber;
   END_REGION

   REGION "ENABLE"
       IF #selStnCount >= 1 THEN

           REGION "SHOW BUTTON DETAILS"
               #animate := #deselected;
           END_REGION

       END_IF;
   END_REGION

   REGION "DISABLE"
       IF #selStnCount = 0 THEN

           REGION "HIDE BUTTON DETAILS"
               #animate := #invisible;
           END_REGION

       END_IF;
   END_REGION

   REGION "APPLY ANIMATION"
       FOR #i := 0 TO #btnCount DO

           REGION "CALCULATE BUTTON POINTER"
               #pBtn := "Pointer Calc: Button Details"(#i);
           END_REGION

           REGION "WHILE Station SELECTED"
               IF #selStnCount <> 0 THEN

                   REGION "COPY TO LOCAL"
                       #btnSelected := #stations.me[#selStnNumber].settings.btnSelection[#pBtn];
                   END_REGION

                   REGION "ANIMATE BUTTON SELECTION

                       REGION "SELECTED"
                           IF #btnSelected THEN
                               #animate := #selected;
                           END_IF;
                       END_REGION

                       REGION "NOT SELECTED"
                           IF NOT #btnSelected THEN
                               #animate := #deselected;
                           END_IF;
                       END_REGION

                   END_REGION

               END_IF;
           END_REGION


           REGION "SEND TO HMI"
               #settings.viewingStation.btns[#i].label.animate := #animate;
               #settings.viewingStation.btns[#i].alloted.animate := #animate;
               #settings.viewingStation.btns[#i].critical.animate := #animate;
               #settings.viewingStation.btns[#i].partNumber.animate := #animate;
           END_REGION

       END_FOR;
   END_REGION
END_FUNCTION

FUNCTION "Populate Station Name" : WString   // FC20, SCL
{ S7_Optimized_Access := 'TRUE' }
VERSION : 0.1
   VAR_INPUT
      line : WString;
      dropZone : USInt;
   END_VAR
BEGIN
   #"Populate Station Name" := CONCAT_WSTRING(IN1 := #line,
                                              IN2 := wstring#' ',
                                              IN3 := "Strip Sign"(USINT_TO_WSTRING(#dropZone)));
END_FUNCTION

FUNCTION "Pointer Calc: Button Details" : Int   // FC21, SCL
{ S7_Optimized_Access := 'TRUE' }
VERSION : 0.1
   VAR_INPUT
      index : Int;
   END_VAR
   VAR_TEMP
      val : Int;
   END_VAR
BEGIN
   IF #index MOD 2 = 0 THEN
       #val := 7 - #index / 2;
   END_IF;

   IF #index MOD 2 <> 0 THEN
       #val := 3 - #index / 2;
   END_IF;

   #"Pointer Calc: Button Details" := #val;
END_FUNCTION

FUNCTION "Buffer Part Req Log Row: Generate" : "Part Req Log Row"   // FC22, SCL
{ S7_Optimized_Access := 'TRUE' }
VERSION : 0.1
   VAR_INPUT
      address : Int;
      "type" : Int;
   END_VAR
   VAR_TEMP
      retVal : Int;
   END_VAR
BEGIN
   REGION "ADDRESS"
       #"Buffer Part Req Log Row: Generate".address := #address;
   END_REGION

   REGION "REQUEST TYPE"
       #"Buffer Part Req Log Row: Generate".reqType := #type;
   END_REGION

   REGION "TIME STAMP"
       #retVal := RD_SYS_T(#"Buffer Part Req Log Row: Generate".timeStamp);
   END_REGION
END_FUNCTION

FUNCTION "Sim to Global" : Void   // FC23, SCL
{ S7_Optimized_Access := 'TRUE' }
VERSION : 0.1
   VAR_INPUT
      simStations : "Simulated Stations";
   END_VAR
   VAR_IN_OUT
      stations : "Stations";
   END_VAR
   VAR_TEMP
      btnCount : Int;
      firstStn : Int;
      i : Int;
      j : Int;
      pSim : Int;
      pStn : Int;
      simKP8Count : Int;
      stnCount : Int;
   END_VAR
BEGIN
   REGION "COPY TO LOCAL"
       #btnCount := "ptsPerStn";
       #firstStn := #simStations.firstStn;
       #simKP8Count := "simKP8Count";
       #stnCount := "stnCount";
   END_REGION

   REGION "FOR EACH STATION"
       FOR #i := 0 TO #simKP8Count DO

           REGION "CALCULATE POINTER"
               #pStn := #i + #firstStn;
               #pSim := #i;
           END_REGION

           REGION "UPPER LIMIT ROLL OVER"
               IF #pStn > #stnCount THEN
                   #pStn := #firstStn + #i - #stnCount - 1;
               END_IF;
           END_REGION

           REGION "COPY SIMULATED PRESSES"
               #stations.me[#pStn].kp8In := #simStations.me[#pSim].btn.actuate;
           END_REGION

       END_FOR;
   END_REGION
END_FUNCTION

FUNCTION "Pointer Calc: KP8 Labels" : Int   // FC25, SCL
{ S7_Optimized_Access := 'TRUE' }
VERSION : 0.1
   VAR_INPUT
      index : Int;
   END_VAR
   VAR_TEMP
      val : Int;
   END_VAR
BEGIN
   IF #index >= 4 THEN
       #val := 7 - (#index - 4) * 2;
   END_IF;

   IF #index <= 3 THEN
       #val := 8 - #index * 2;
   END_IF;

   #"Pointer Calc: KP8 Labels" := #val;
END_FUNCTION

FUNCTION "KP8 Color to Sim Animation" : USInt   // FC26, SCL
{ S7_Optimized_Access := 'TRUE' }
VERSION : 0.1
   VAR_INPUT
      kp8Color : DWord;
      btnNumber : Int;
   END_VAR
   VAR_TEMP
      animate : USInt;
      blue : USInt;
      colorDWord : DWord;
      colorInt : DInt;
      green : USInt;
      off : USInt;
      red : USInt;
      white : USInt;
      yellow : USInt;
   END_VAR
   VAR CONSTANT
      blueMask : DInt := 16#0000_0100;
      btnMask : DInt := 16#0101_0100;
      greenMask : DInt := 16#0001_0000;
      offMask : DInt := 16#0000_0000;
      redMask : DInt := 16#0100_0000;
      whiteMask : DInt := 16#0101_0100;
      yellowMask : DInt := 16#0101_0000;
   END_VAR
BEGIN
   REGION "COPY TO LOCAL"
       #blue := "BgLBl";
       #green := "BgLGr";
       #off := "BgGray";
       #red := "BgLRd";
       #white := "BgWh";
       #yellow := "BgLYe";
   END_REGION

   REGION "ISOLATE BUTTON COLOR"
       #colorDWord := SHR_DWORD(IN := #kp8Color,N := INT_TO_ULINT(#btnNumber));
       #colorDWord := #colorDWord AND #btnMask;
       #colorInt := DWORD_TO_DINT(#colorDWord);
   END_REGION

   REGION "DETERMINE ANIMATION"
       CASE #colorInt OF
           #blueMask:
               #animate := #blue;
           #greenMask:
               #animate := #green;
           #redMask:
               #animate := #red;
           #whiteMask:
               #animate := #white;
           #yellowMask:
               #animate := #yellow;
           ELSE
               #animate := #off;
       END_CASE;
   END_REGION

   REGION "RETURN VALUE"
       #"KP8 Color to Sim Animation" := #animate;
   END_REGION
END_FUNCTION

FUNCTION "Word Wrap" : WString   // FC28, SCL
{ S7_Optimized_Access := 'TRUE' }
VERSION : 0.1
   VAR_INPUT
      stringIn : WString;
      maxLength : Int;
   END_VAR
   VAR_TEMP
      length : Int;
      charBox : Array[0.."lStringLen"] of WChar;
      stringBox : Array[0.."lStringLen"] of WString["lStringLen"];
      count : UInt;
      status : Int;
      i : Int;
      pStringBox : Int;
      output : WString;
      savedOutput : WString;
      lineBox : Array[0..10] of WString["lStringLen"];
      pLineBox : Int;
      lengthTest : WString;
   END_VAR
   VAR CONSTANT
      space : WString := WSTRING#' ';
      blank : WString;
      lineBreak : WString := WSTRING#'$L';
   END_VAR
BEGIN
   #length := LEN(#stringIn);

   IF #length <= #maxLength THEN
       #output := #stringIn;
   END_IF;

   IF #length > #maxLength THEN

       Strg_TO_Chars(
                     Strg := #stringIn,
                     pChars := 0,
                     Cnt => #count,
                     Chars := #charBox
       );

       FOR #i := 0 TO "lStringLen" DO

           IF #charBox[#i] = #space THEN
               IF #charBox[#i + 1] = #space THEN
                   EXIT;
               END_IF;
           END_IF;

           IF #i = 0 THEN
               #stringBox[#pStringBox] := #charBox[#i];
           END_IF;

           IF #i >= 1 THEN
               #stringBox[#pStringBox] := CONCAT_WSTRING(IN1 := #stringBox[#pStringBox],
                                                         IN2 := #charBox[#i]);
           END_IF;

           IF #charBox[#i] = #space THEN
               #stringBox[#pStringBox] := "Trim"(#stringBox[#pStringBox]);
               #pStringBox := #pStringBox + 1;
           END_IF;

           IF #charBox[#i] = #lineBreak THEN
               #stringBox[#pStringBox] := LEFT(IN := #stringBox[#pStringBox],
                                               L := LEN(#stringBox[#pStringBox]) - 1);
               #pStringBox := #pStringBox + 1;
               #stringBox[#pStringBox] := #lineBreak;
               #pStringBox := #pStringBox + 1;
           END_IF;

       END_FOR;


       FOR #i := 0 TO "lStringLen" DO

           IF #stringBox[#i] = #blank THEN
               IF #stringBox[#i + 1] = #blank THEN
                   #lineBox[#pLineBox] := "Trim"(#lineBox[#pLineBox]);
                   EXIT;
               END_IF;
           END_IF;

           IF #stringBox[#i] = #lineBreak THEN
               #lineBox[#pLineBox] := "Trim"(#lineBox[#pLineBox]);
               #pLineBox := #pLineBox + 1;
               #lineBox[#pLineBox] := #lineBreak;
               #pLineBox := #pLineBox + 1;
           END_IF;


           IF #stringBox[#i] <> #lineBreak THEN

               IF #i = 0 THEN
                   #lengthTest := #stringBox[#i];
               END_IF;

               IF #i >= 1 THEN
                   #lengthTest := CONCAT_WSTRING(IN1 := #lineBox[#pLineBox],
                                                 IN2 := #space,
                                                 IN3 := #stringBox[#i]);
               END_IF;

               IF LEN(#lengthTest) <= #maxLength THEN
                   #lineBox[#pLineBox] := #lengthTest;
               END_IF;

               IF LEN(#lengthTest) > #maxLength THEN
                   #lineBox[#pLineBox] := "Trim"(#lineBox[#pLineBox]);
                   #lineBox[#pLineBox] := "Trim"(#lineBox[#pLineBox]);
                   #pLineBox := #pLineBox + 1;
                   #lineBox[#pLineBox] := #stringBox[#i];
               END_IF;
           END_IF;

       END_FOR;

       FOR #i := 0 TO 10 DO

           IF #lineBox[#i] = #space OR #lineBox[#i] = WString#'' THEN
               EXIT;
           END_IF;
           IF #i = 0 THEN
               #output := #lineBox[#i];
           END_IF;
           IF #i >= 1 THEN
               IF #lineBox[#i] = #lineBreak THEN
                   #output := #output;
               END_IF;
               IF #lineBox[#i] <> #lineBreak THEN
                   #output := CONCAT_WSTRING(IN1 := #output,
                                             IN2 := #lineBreak,
                                             IN3 := #lineBox[#i]);
               END_IF;
           END_IF;

       END_FOR;

       #output := "Trim"(#output);

   END_IF;

   #"Word Wrap" := #output;
END_FUNCTION

FUNCTION "Trim" : WString   // FC29, SCL
{ S7_Optimized_Access := 'TRUE' }
VERSION : 0.1
   VAR_INPUT
      stringIn : WString;
   END_VAR
   VAR_TEMP
      output : WString;
   END_VAR
   VAR CONSTANT
      space : WString := WSTRING#' ';
   END_VAR
BEGIN
   #output := #stringIn;
   IF LEFT(IN := #output, L := 1) = #space THEN
       #output := RIGHT(IN := #output, L := LEN(#output) - 1);
   END_IF;
   IF RIGHT(IN := #output, L := 1) = #space THEN
       #output := LEFT(IN := #output, L := LEN(#output) - 1);
   END_IF;
   #Trim := #output;
END_FUNCTION

FUNCTION "Recipe Select Button" : Void   // FC31, SCL
{ S7_Optimized_Access := 'TRUE' }
VERSION : 0.1
   VAR_INPUT
      visRows : Int;
      lib : "Menu: Library";
      actuate : Bool;
      maxRows : Int;
      btnNum : Int;
   END_VAR
   VAR_IN_OUT
      recipeSelectScreen : "HSS: Menu Selection Screen";
   END_VAR
   VAR_TEMP
      eval : "HSS: Menu Selection Screen";
      pRowVisLbl : Int;
      pRowInvisLbl : Int;
      pRowTxt : Int;
      pRecipeTxt : Int;
      maxLen : Int;
   END_VAR
BEGIN
   #eval := #recipeSelectScreen;

   REGION "NARROW"
       IF #maxRows > #visRows THEN
           #pRowVisLbl := #btnNum + #visRows;
           #pRowInvisLbl := #btnNum + (3 * #visRows);
           #maxLen := 22;
       END_IF;
   END_REGION


   REGION "WIDE"
       IF #maxRows <= #visRows THEN
           #pRowVisLbl := #btnNum + (3 * #visRows);
           #pRowInvisLbl := #btnNum + #visRows + 1;
           #maxLen := 28;
       END_IF;
   END_REGION


   REGION "ROW COUNT INDEPENDENT"
       #pRowTxt := (#btnNum * 2) + #visRows;
       #pRecipeTxt := #pRowTxt + 1;
   END_REGION


   REGION "DRAW"
       #eval.animate[#pRowVisLbl] := "BgGray";
       #eval.animate[#pRowInvisLbl] := "invisible";
       #eval.txt[#pRowTxt] := "Strip Sign"(DINT_TO_WSTRING(#btnNum));
       #eval.txt[#pRecipeTxt] := "Word Wrap"(stringIn := #lib.entry[#btnNum],
                                             maxLength := #maxLen);
   END_REGION

   IF #actuate THEN
       #eval.animate[#pRowVisLbl] := "BgLTe";
   END_IF;

   #recipeSelectScreen := #eval;
END_FUNCTION

FUNCTION "Recipe Nav Button" : Void   // FC32, SCL
{ S7_Optimized_Access := 'TRUE' }
VERSION : 0.1
   VAR_INPUT
      visRows : Int;
      actuate : Bool;
      maxRows : Int;
      btnNum : Int;
   END_VAR
   VAR_IN_OUT
      recipeSelectScreen : "HSS: Menu Selection Screen";
   END_VAR
   VAR_TEMP
      eval : "HSS: Menu Selection Screen";
      color : Int;
   END_VAR
BEGIN
   #eval := #recipeSelectScreen;

   REGION "NARROW"
       IF #maxRows > #visRows THEN
           #color := "BgGray";
       END_IF;
   END_REGION


   REGION "WIDE"
       IF #maxRows <= #visRows THEN
           #color := "invisible";
       END_IF;
   END_REGION


   REGION "ROW COUNT INDEPENDENT"
       IF #actuate THEN
           #color := "BgLTe";
       END_IF;
   END_REGION


   REGION "DRAW"
       #eval.animate[#btnNum] := #color;
   END_REGION

   #recipeSelectScreen := #eval;
END_FUNCTION

// ===== library types =====
